            #instTcpSend.REQ := true;
             #instTcpSend.LEN := INT_TO_UDINT(#statSendLenght + 2);

                   IF ((#instTcpSend.DONE)
                       AND (#instTcpSend.BUSY = 0))
                   THEN
                       #instTcpSend.REQ := false;
                       #statStateMQTT := #MQTT_CONNACK;
                       //Delete Send Buffer
                       FOR #statI := 1 TO (#statSendLenght + 2) DO
                           #statSendBuffer[#statI] := 0;
                       END_FOR;
                   ELSIF #instTcpSend.ERROR
                   THEN
                       #statusID := #MQTT_CONNECT;
                       #instTcpSend.REQ := false;
                       #statStateMQTT := #MQTT_ERROR;

                   END_IF;

               END_REGION
               ;
           #MQTT_CONNACK:
               IF #statNewDataRcv THEN

                   IF ((#statRcvBuffer[1] AND b#16#f0) = #MQTT_MSG_TYPE_CONNACK)
                       AND
                       (#statRcvBuffer[4] = #MQTT_CONNACK_ACCEPTED)
                   THEN
                       #statStateMQTT := #MQTT_CONNECTED;
                       #mqttEstablished := true;
                       #busy := false;
                       #statStateMQTTinternal := #IDLE;
                       //start Keep Alive Timer
                       //KeepAliveTImer is set to (Keep Alive (in s) - 2s)
                       #statKeepAliveTime := UINT_TO_TIME((WORD_TO_UINT(#mqttParam.keepAlive) * 1000 - 2000));
                       IF NOT #statKeepAliveOff
                       THEN
                           #statTriggerKeepAlive := true;
                       END_IF;
                       #statNewDataRcv := 0;
                   ELSE
                       #statStateMQTT := #MQTT_ERROR;
                       #statusID := #MQTT_CONNACK;
                   END_IF;
               END_IF;
           #MQTT_CONNECTED:
               IF #publish
                   AND NOT #statPublishOld
                   AND (#statStateMQTTinternal=#IDLE)
               THEN
                   #statStateMQTTinternal := #MQTT_PUBLISH;
                   #published := 0;
                   #error := 0;
                  #statTriggerKeepAlive := false;
                   #statPacketID := #statPacketID + 1;
               END_IF;
               #statPublishOld := #publish;

                IF (#instKeepAlive.Q)
                    AND (#statStateMQTTinternal = #IDLE)
                    AND (NOT #statKeepAliveOff)
                THEN
                    #statStateMQTTinternal := #MQTT_PING;
                    #statTriggerKeepAlive := false;
                END_IF;
                CASE #statStateMQTTinternal OF
                    #IDLE:
                        #published := 0;
                        ;
                    #MQTT_PUBLISH:
                        ;
                        #busy := true;
                        #statConnectLenghtOffset := 0;
                        #statConnectLenght := LEN(IN := #mqttParam.topic) + LEN(IN := #mqttParam.message) + 2;
                        #statSendBuffer[1] := 16#30;
                        #statSendBuffer[1].%X0 := #mqttParam.publishFlag.retain;
                        #statSendBuffer[1].%X3 := false;
                        CASE #mqttParam.publishFlag.qualityOfService OF
                            0:
                                #statSendBuffer[1].%X1 := 0;
                                #statSendBuffer[1].%X2 := 0;
                            1:
                                #statSendBuffer[1].%X1 := 1;
                                #statSendBuffer[1].%X2 := 0;
                                //2 Byte Packet Identifiert added
                                #statConnectLenght := #statConnectLenght + 2;
                            2:
                                #statSendBuffer[1].%X1 := 0;
                                #statSendBuffer[1].%X2 := 1;
                                //2 Byte Packet Identifiert added
                                #statConnectLenght := #statConnectLenght + 2;
                            ELSE:
                                ;
                                #statStateMQTT := #MQTT_ERROR;
                                #statusID := #MQTT_PUBLISH;
                        END_CASE;
                        #statSendLenght := #statConnectLenght;
                        WHILE (#statConnectLenght > 0)
                        DO
                            #statConnectEncodedLenght := #statConnectLenght MOD 128;
                            #statConnectLenght := #statConnectLenght / 128;
                            // if there are more data to encode, set the top bit of this byte
                            IF #statConnectLenght > 0
                            THEN
                                #statConnectEncodedLenght := #statConnectEncodedLenght OR 128;
                                #statSendBuffer[2 + #statConnectLenghtOffset] := INT_TO_BYTE(#statConnectEncodedLenght);
                                #statConnectLenghtOffset := #statConnectLenghtOffset + 1;
                            ELSE
                                #statSendBuffer[2 + #statConnectLenghtOffset] := INT_TO_BYTE(#statConnectEncodedLenght);
                            END_IF;
                        END_WHILE;
                        #statSendLenght := #statSendLenght + #statConnectLenghtOffset;
                        //Variable Header
                        #tempLenght := INT_TO_WORD(LEN(IN := #mqttParam.topic));
                        #statSendBuffer[3 + #statConnectLenghtOffset] := #tempLenght.%B1;
                        #statSendBuffer[4 + #statConnectLenghtOffset] := #tempLenght.%B0;
                        Strg_TO_Chars(Strg := #mqttParam.topic,
                                      pChars := 0,
                                      Cnt => #tempCountChars,
                                      Chars := #tempStringToChar);
                        FOR #statI := 0 TO UINT_TO_INT(#tempCountChars - 1) DO
                            #statSendBuffer[5 + #statConnectLenghtOffset + #statI] := #tempStringToChar[#statI];
                        END_FOR;
                        #statConnectLenghtOffset := #statConnectLenghtOffset + #statI;
                        IF (#mqttParam.publishFlag.qualityOfService > 0)
                        THEN

                            #statSendBuffer[5 + #statConnectLenghtOffset] := #statPacketID.%B1;
                            #statSendBuffer[6 + #statConnectLenghtOffset] := #statPacketID.%B0;
                            //Payload
                            Strg_TO_Chars(Strg := #mqttParam.message,
                                          pChars := 0,
                                          Cnt => #tempCountChars,
                                          Chars := #tempStringToChar);
                            FOR #statI := 0 TO UINT_TO_INT(#tempCountChars - 1) DO
                                #statSendBuffer[7 + #statConnectLenghtOffset + #statI] := #tempStringToChar[#statI];
                            END_FOR;
                            #instTcpSend.LEN := INT_TO_UDINT(#statSendLenght + 2);
                        ELSE
                            Strg_TO_Chars(Strg := #mqttParam.message,
                                          pChars := 0,
                                          Cnt => #tempCountChars,
                                          Chars := #tempStringToChar);
                            FOR #statI := 0 TO UINT_TO_INT(#tempCountChars - 1) DO
                                #statSendBuffer[5 + #statConnectLenghtOffset + #statI] := #tempStringToChar[#statI];
                            END_FOR;
                            #instTcpSend.LEN := INT_TO_UDINT(#statSendLenght + 2);
                        END_IF;

                        #instTcpSend.REQ := true;


                        IF ((#instTcpSend.DONE)
                            AND (#instTcpSend.BUSY = 0))
                        THEN
                            #instTcpSend.REQ := false;
                            IF (#mqttParam.publishFlag.qualityOfService > 0)
                            THEN
                                #statPacketIDAck := #statPacketID;
                                #statStateMQTTinternal := #MQTT_PUBACK;
                            ELSE
                                //QoS = 0; finish here
                                #published := true;
                                #busy := false;
                                #statNewDataRcv := false;
                                IF NOT #statKeepAliveOff
                                THEN
                                    #statTriggerKeepAlive := true;
                                END_IF;

                                #statStateMQTTinternal := #IDLE;
                            END_IF;
                        ELSIF #instTcpSend.ERROR
                        THEN
                            #statusID := #MQTT_PUBLISH;
                            #instTcpSend.REQ := false;
                            #statStateMQTT := #MQTT_ERROR;
                            #status := #instTcpSend.STATUS;
                        END_IF;
                    #MQTT_PUBACK:
                        IF #statNewDataRcv THEN
                            IF ((#statRcvBuffer[1] AND b#16#f0) = #MQTT_MSG_TYPE_PUBACK)
                                OR
                                ((#statRcvBuffer[1] AND b#16#f0) = INT_TO_WORD(#MQTT_MSG_TYPE_PUBREC))
                            THEN
                                IF
                                    (#statRcvBuffer[3] = #statPacketIDAck.%B1)
                                    AND
                                    (#statRcvBuffer[4] = #statPacketIDAck.%B0)
                                THEN
                                    IF (#mqttParam.publishFlag.qualityOfService = 1)
                                    THEN
                                        //QoS = 1; finish here
                                        #statStateMQTTinternal := #MQTT_IDLE;
                                        #published := true;
                                        #busy := false;
                                        #statNewDataRcv := false;
                                        //Re-Activate Kepp Alive Timer
                                        IF NOT #statKeepAliveOff
                                        THEN
                                            #statTriggerKeepAlive := true;
                                        END_IF;

                                        #statStateMQTTinternal := #IDLE;
                                    ELSE
                                        #statStateMQTTinternal := #MQTT_PUBREL;
                                    END_IF;
                                ELSE
                                    #statNewDataRcv := false;
                                END_IF;
                            ELSE
                                #statStateMQTT := #MQTT_ERROR;
                                #statusID := #MQTT_PUBACK;
                            END_IF;
                        END_IF;
                    #MQTT_PUBREL:
                        //fixed Header
                        #statSendBuffer[1] := 16#62;
                        #statSendBuffer[2] := 2;
                        //Variable Header
                        #statSendBuffer[3] := #statPacketID.%B1;
                        #statSendBuffer[4] := #statPacketID.%B0;
                        #instTcpSend.LEN := INT_TO_UDINT(4);
                        #instTcpSend.REQ := true;

                        IF ((#instTcpSend.DONE)
                            AND (#instTcpSend.BUSY = 0))
                        THEN
                            #instTcpSend.REQ := false;
                            #statPacketIDAck := #statPacketID;
                            #statStateMQTTinternal := #MQTT_PUBCOMP;

                        ELSIF #instTcpSend.ERROR
                        THEN
                            #statusID := #MQTT_PUBREL;
                            #instTcpSend.REQ := false;
                            #statStateMQTT := #MQTT_ERROR;
                            #status := #instTcpSend.STATUS;
                        END_IF;
                    #MQTT_PUBCOMP:
                        IF #statNewDataRcv THEN
                            IF ((#statRcvBuffer[1] AND b#16#f0) = #MQTT_MSG_TYPE_PUBCOM)
                            THEN
                                IF
                                    (#statRcvBuffer[3] = #statPacketIDAck.%B1)
                                    AND
                                    (#statRcvBuffer[4] = #statPacketIDAck.%B0)
                                THEN
                                    //QoS = 2; finish here
                                    #statStateMQTTinternal := #MQTT_IDLE;
                                    #published := true;
                                    #busy := false;
                                    #statNewDataRcv := false;
                                    //Re-Activate Kepp Alive Timer
                                    IF NOT #statKeepAliveOff
                                    THEN
                                        #statTriggerKeepAlive := true;
                                    END_IF;

                                    #statStateMQTTinternal := #IDLE;
                                ELSE
                                    #statStateMQTT := #MQTT_ERROR;
                                    #statusID := #MQTT_PUBCOMP;
                                END_IF;
                            END_IF;
                        END_IF;
                    #MQTT_PING:

                        #busy := true;
                        //Build fixed Header
                        //Message Type
                        #statSendBuffer[1] := INT_TO_BYTE(#MQTT_MSG_TYPE_PING);
                        //Remaining Lenght (must be O)
                        #statSendBuffer[2] := 0;
                        #instTcpSend.REQ := true;
                        #instTcpSend.LEN := 2;

                        IF ((#instTcpSend.DONE)
                            AND (#instTcpSend.BUSY = 0))
                        THEN
                            #instTcpSend.REQ := false;
                            #statStateMQTTinternal := #MQTT_PINGRESP;
                        ELSIF #instTcpSend.ERROR
                        THEN
                            #statusID := #MQTT_PING;
                            #instTcpSend.REQ := false;
                            #statStateMQTT := #MQTT_ERROR;
                            #status := #instTcpSend.STATUS;
                        END_IF;
                    #MQTT_PINGRESP:
                        IF #statNewDataRcv
                        THEN
                            IF ((#statRcvBuffer[1] AND b#16#f0) = #MQTT_MSG_TYPE_PINGRESP)
                            THEN
                                #busy := false;
                                #statNewDataRcv := false;
                                #statTriggerKeepAlive := true;
                                #statStateMQTTinternal := #IDLE;
                            END_IF;
                        ELSE
                            #statNewDataRcv := false;
                        END_IF;

                END_CASE;
           #MQTT_DISCONNECT:
           #busy := 0;
           //Build fixed Header
           //Message Type
           #statSendBuffer[1] := INT_TO_BYTE(#MQTT_MSG_TYPE_DISCONNECT);
           //Remaining Lenght (must be O)
           #statSendBuffer[2] := 0;
           #instTcpSend.REQ := true;
           #instTcpSend.LEN := 2;

           IF ((#instTcpSend.DONE)
               AND (#instTcpSend.BUSY = 0))
           THEN
               IF NOT #enable THEN
                   #statStateTCP := #TCP_DISCONNECT;
               END_IF;
               #instTcpSend.REQ := false;
               #statStateMQTT := #MQTT_DISCONNECTED;
               #statStateMQTTinternal := #IDLE;
           ELSIF #instTcpSend.ERROR
           THEN
               IF NOT #enable THEN
                   #statStateTCP := #TCP_DISCONNECT;
               END_IF;
               #statusID := #MQTT_DISCONNECT;
               #instTcpSend.REQ := false;
               #statStateMQTT := #MQTT_ERROR;
               #status := #instTcpSend.STATUS;
           END_IF;
               #MQTT_ERROR:

               REGION Errorhandling MQTT
                   #error := true;
                   #busy := false;
                   #statStateMQTTinternal := #IDLE;
                   #statTriggerKeepAlive := 0;
                   #statKeepAliveOff := false;
                 CASE #statusID OF
                     #MQTT_CONNECT_FLAG_CHECK:
                         #mqttEstablished := false;
                         #statStateMQTT := #MQTT_DISCONNECTED;
                         ;
                     #MQTT_CONNECT:
                         #mqttEstablished := false;
                         #status := #instTcpSend.STATUS;   ;
                         #statStateMQTT := #MQTT_DISCONNECTED;
                       #MQTT_CONNACK:
                           #mqttEstablished := false;
                           #status := #statRcvBuffer[4];
                           #statStateMQTT := #MQTT_DISCONNECTED;
                       #MQTT_PUBLISH:
                               #published := false;
                               #statStateMQTT := #MQTT_CONNECTED;
                               #MQTT_PUBACK,#MQTT_PUBCOMP,#MQTT_PUBREL:
                           #published := false;
                           #status :=#MQTT_ERROR_PACKETID;
                           #statStateMQTT := #MQTT_CONNECTED;
                       #MQTT_PINGRESP:;
                           #MQTT_PING:;
                       #MQTT_DISCONNECT:
                           #mqttEstablished := false;
                          ;
                       ELSE
                           ;
                   END_CASE;
              END_REGION
               ;



       END_CASE
       ;
END_FUNCTION_BLOCK

FUNCTION_BLOCK "FB_MQTT"   // FB5, LAD
{ S7_Optimized_Access := 'TRUE' }
VERSION : 0.1
BEGIN
END_FUNCTION_BLOCK

FUNCTION_BLOCK "FB_concatScrings"   // FB6, LAD
{ S7_Optimized_Access := 'TRUE' }
VERSION : 0.1
   VAR_INPUT
      temperature1 : Real;
      temperature2 : Real;
      temperature3 : Real;
      temperature4 : Real;
      rtd_ch0 : Real;
      rtd_ch1 : Real;
      rtd_ch2 : Real;
      rtd_ch3 : Real;
      presaCounter : UDInt;
      PresaHitrost : Int;
      PresaisRunning : Int;
   END_VAR
   VAR_OUTPUT
      strCombinedString : String;
   END_VAR
   VAR
      tempStr1 : String;
      tempStr2 : String;
      tempStr3 : String;
      tempStr4 : String;
      counterStr : String;
      isRunningStr : String;
      currentSpeedStr : String;
      combinedStr : String;
      rtdStr0 : String;
      rtdStr1 : String;
      rtdStr2 : String;
      rtdStr3 : String;
   END_VAR
BEGIN

REGION Network 2 (SCL)
   // Convert REAL values to STRING
   // 
    VAL_STRG(IN:=#temperature1,
              SIZE:=10,
              PREC:=4,
              FORMAT:=0000,
              P:=16,
              OUT=>#tempStr1);

   //#tempStr1 := REAL_TO_STRING(#temperature1);

     VAL_STRG(IN := #temperature2,
              SIZE := 10,
              PREC := 4,
              FORMAT := 0000,
              P := 16,
              OUT => #tempStr2);

     VAL_STRG(IN := #temperature3,
              SIZE := 10,
              PREC := 4,
              FORMAT := 0000,
              P := 16,
              OUT => #tempStr3);

     VAL_STRG(IN := #temperature4,
              SIZE := 10,
              PREC := 4,
              FORMAT := 0000,
              P := 16,
              OUT => #tempStr4);

   //convert RTD inputs to string
   // Convert RTD values to STRING
   VAL_STRG(IN := #rtd_ch0,
            SIZE := 10,
            PREC := 4,
            FORMAT := 0000,
            P := 16,
            OUT => #rtdStr0);
   VAL_STRG(IN := #rtd_ch1,
            SIZE := 10,
            PREC := 4,
            FORMAT := 0000,
            P := 16,
            OUT => #rtdStr1);
   VAL_STRG(IN := #rtd_ch2,
            SIZE := 10,
            PREC := 4,
            FORMAT := 0000,
            P := 16,
            OUT => #rtdStr2);
   VAL_STRG(IN := #rtd_ch3,
            SIZE := 10,
            PREC := 4,
            FORMAT := 0000,
            P := 16,
            OUT => #rtdStr3);

   // convert int to string
     #currentSpeedStr := ' ';
     VAL_STRG(IN := #PresaHitrost,
              SIZE := 3,
              PREC := 0,
              FORMAT := 0000,
              P := 1,
              OUT => #currentSpeedStr);


   // Convert DINT to STRING
   #counterStr := '';
   VAL_STRG(IN := #presaCounter,
            SIZE := 5,
            PREC := 0,
            FORMAT := 0000,
            P := 1,
            OUT => #counterStr);

   // Convert BOOL to STRING (represent TRUE/FALSE)
   IF #PresaisRunning = 1 THEN
       #isRunningStr := '1';
   ELSE
       #isRunningStr := '0';
   END_IF;

   // Combine all strings into a JSON format
   #combinedStr := '{';
   #combinedStr := CONCAT(IN1 := #combinedStr, IN2 := '"temperature1":');
   #combinedStr := CONCAT(IN1 := #combinedStr, IN2 := #tempStr1);
   #combinedStr := CONCAT(IN1 := #combinedStr, IN2 := ',');
   #combinedStr := CONCAT(IN1 := #combinedStr, IN2 := '"temperature2":');
   #combinedStr := CONCAT(IN1 := #combinedStr, IN2 := #tempStr2);
   #combinedStr := CONCAT(IN1 := #combinedStr, IN2 := ',');
   #combinedStr := CONCAT(IN1 := #combinedStr, IN2 := '"temperature3":');
   #combinedStr := CONCAT(IN1 := #combinedStr, IN2 := #tempStr3);
   #combinedStr := CONCAT(IN1 := #combinedStr, IN2 := ',');
   #combinedStr := CONCAT(IN1 := #combinedStr, IN2 := '"temperature4":');
   #combinedStr := CONCAT(IN1 := #combinedStr, IN2 := #tempStr4);
   #combinedStr := CONCAT(IN1 := #combinedStr, IN2 := ',');

   (* #combinedStr := CONCAT(IN1 := #combinedStr, IN2 := '"rtd_ch0":');
   #combinedStr := CONCAT(IN1 := #combinedStr, IN2 := #rtdStr0);
   #combinedStr := CONCAT(IN1 := #combinedStr, IN2 := ',');

   #combinedStr := CONCAT(IN1 := #combinedStr, IN2 := '"rtd_ch1":');
   #combinedStr := CONCAT(IN1 := #combinedStr, IN2 := #rtdStr1);
   #combinedStr := CONCAT(IN1 := #combinedStr, IN2 := ',');
   *)
   #combinedStr := CONCAT(IN1 := #combinedStr, IN2 := '"rtd_ch2":');
   #combinedStr := CONCAT(IN1 := #combinedStr, IN2 := #rtdStr2);
   #combinedStr := CONCAT(IN1 := #combinedStr, IN2 := ',');


   #combinedStr := CONCAT(IN1 := #combinedStr, IN2 := '"counter":');
   #combinedStr := CONCAT(IN1 := #combinedStr, IN2 := #counterStr);
   #combinedStr := CONCAT(IN1 := #combinedStr, IN2 := ',');
   #combinedStr := CONCAT(IN1 := #combinedStr, IN2 := '"isRunning":');
   #combinedStr := CONCAT(IN1 := #combinedStr, IN2 := #isRunningStr);
   #combinedStr := CONCAT(IN1 := #combinedStr, IN2 := ',');
   #combinedStr := CONCAT(IN1 := #combinedStr, IN2 := '"currentSpeed":');
   #combinedStr := CONCAT(IN1 := #combinedStr, IN2 := #currentSpeedStr);
   #combinedStr := CONCAT(IN1 := #combinedStr, IN2 := '}');

   // Now combinedStr contains the concatenated string in JSON format
   #strCombinedString := #combinedStr;
END_REGION
END_FUNCTION_BLOCK

FUNCTION_BLOCK "FB_CONCAT_STRINGS_FOR_MQTT"   // FB7, LAD
{ S7_Optimized_Access := 'TRUE' }
VERSION : 0.1
   VAR_INPUT
      temperature1 : Real;
      temperature2 : Real;
      temperature3 : Real;
      temperature4 : Real;
   END_VAR
   VAR_OUTPUT
      strCombinedString : String;
      q_aStringToSendToMqtt : Array[0..1] of String;
   END_VAR
   VAR
      tempStr1 : String;
      tempStr2 : String;
      tempStr3 : String;
      tempStr4 : String;
      combinedStr : String;
      lenghtOfCombinedString : Int;
      Static_1 : Int;
      assocValues : Array[0..3] of DInt;
      combineStr_1 : String;
      combineStr_2 : String;
   END_VAR
BEGIN

REGION Network 2 (SCL)
   // Convert REAL values to STRING
   // 
   VAL_STRG(IN := #temperature1,
            SIZE := 10,
            PREC := 4,
            FORMAT := 0000,
            P := 16,
            OUT => #tempStr1);

   //#tempStr1 := REAL_TO_STRING(#temperature1);

   VAL_STRG(IN := #temperature2,
            SIZE := 10,
            PREC := 4,
            FORMAT := 0000,
            P := 16,
            OUT => #tempStr2);

   VAL_STRG(IN := #temperature3,
            SIZE := 10,
            PREC := 4,
            FORMAT := 0000,
            P := 16,
            OUT => #tempStr3);

   VAL_STRG(IN := #temperature4,
            SIZE := 10,
            PREC := 4,
            FORMAT := 0000,
            P := 16,
            OUT => #tempStr4);


   // Combine all strings into a JSON format
   #combinedStr := '{';
   #combinedStr := CONCAT(IN1 := #combinedStr, IN2 := '"temperature1":');
   #combinedStr := CONCAT(IN1 := #combinedStr, IN2 := #tempStr1);
   #combinedStr := CONCAT(IN1 := #combinedStr, IN2 := ',');
   #combinedStr := CONCAT(IN1 := #combinedStr, IN2 := '"temperature2":');
   #combinedStr := CONCAT(IN1 := #combinedStr, IN2 := #tempStr2);
   #combinedStr := CONCAT(IN1 := #combinedStr, IN2 := ',');
   #combinedStr := CONCAT(IN1 := #combinedStr, IN2 := '"temperature3":');
   #combinedStr := CONCAT(IN1 := #combinedStr, IN2 := #tempStr3);
   #combinedStr := CONCAT(IN1 := #combinedStr, IN2 := ',');
   #combinedStr := CONCAT(IN1 := #combinedStr, IN2 := '"temperature4":');
   #combinedStr := CONCAT(IN1 := #combinedStr, IN2 := #tempStr4);
   #combinedStr := CONCAT(IN1 := #combinedStr, IN2 := '}');

   // Now combinedStr contains the concatenated string in JSON format
   #strCombinedString := #combinedStr;

   #lenghtOfCombinedString := LEN(#combinedStr);


   // Check if the length exceeds 254 characters
   IF #lenghtOfCombinedString > 254 THEN
       // Extract the first 254 characters for combineStr_1
       #combineStr_1 := LEFT(IN := #combinedStr, L := 254);

       // Extract the remaining characters for combineStr_2
       #combineStr_2 := RIGHT(IN := #combinedStr, L := #lenghtOfCombinedString - 254);
   ELSE
       // If length is less than or equal to 254, use the entire string in combineStr_1
       #combineStr_1 := #combinedStr;
       #combineStr_2 := '';  // Set combineStr_2 to an empty string
   END_IF;

   #q_aStringToSendToMqtt[0] := #combineStr_1;
   #q_aStringToSendToMqtt[1] := #combineStr_2;
END_REGION
END_FUNCTION_BLOCK

FUNCTION_BLOCK "FB_CONCAT_STRINGS_FOR_MQTT_1"   // FB9, LAD
{ S7_Optimized_Access := 'TRUE' }
VERSION : 0.1
   VAR_INPUT
      temperature1 : Real;
      temperature2 : Real;
      temperature3 : Real;
      temperature4 : Real;
      customText : String;
   END_VAR
   VAR_OUTPUT
      strCombinedString : String;
      q_aStringToSendToMqtt : Array[0..1] of String;
   END_VAR
   VAR
      tempStr1 : String;
      tempStr2 : String;
      tempStr3 : String;
      tempStr4 : String;
      combinedStr : String;
      lenghtOfCombinedString : Int;
      Static_1 : Int;
      assocValues : Array[0..3] of DInt;
      combineStr_1 : String;
      combineStr_2 : String;
      currentStrLength : Int;
      tempStrLength : Int;
      SafeConcat : "FB_saveConcat";
   END_VAR
BEGIN

REGION Network 2 (SCL)
   // Initialize variables
   #combinedStr := '{';
   #combineStr_1 := ''; // First part of the JSON
   #combineStr_2 := ''; // Second part of the JSON

   // Convert REAL values to STRING
   VAL_STRG(IN := #temperature1,
            SIZE := 10,
            PREC := 4,
            FORMAT := 0000,
            P := 16,
            OUT => #tempStr1);

   VAL_STRG(IN := #temperature2,
            SIZE := 10,
            PREC := 4,
            FORMAT := 0000,
            P := 16,
            OUT => #tempStr2);

   VAL_STRG(IN := #temperature3,
            SIZE := 10,
            PREC := 4,
            FORMAT := 0000,
            P := 16,
            OUT => #tempStr3);

   VAL_STRG(IN := #temperature4,
            SIZE := 10,
            PREC := 4,
            FORMAT := 0000,
            P := 16,
            OUT => #tempStr4);

   // Start constructing the JSON string

   // Concatenate temperature1
   #SafeConcat(IN1 := #customText,
               IN2 := #tempStr1,
               combineStr_1 := #combineStr_1,
               combineStr_2 := #combineStr_2,
               SafeConcat => #combinedStr);

   #SafeConcat(IN1 := ',',
               IN2 := '',
               combineStr_1 := #combineStr_1,
               combineStr_2 := #combineStr_2,
               SafeConcat => #combinedStr);

   // Concatenate temperature2
   #SafeConcat(IN1 := '"temperature2":',
               IN2 := #tempStr2,
               combineStr_1 := #combineStr_1,
               combineStr_2 := #combineStr_2,
               SafeConcat => #combinedStr);

   #SafeConcat(IN1 := ',',
               IN2 := '',
               combineStr_1 := #combineStr_1,
               combineStr_2 := #combineStr_2,
               SafeConcat => #combinedStr);

   // Concatenate temperature3
   #SafeConcat(IN1 := '"temperature3":',
               IN2 := #tempStr3,
               combineStr_1 := #combineStr_1,
               combineStr_2 := #combineStr_2,
               SafeConcat => #combinedStr);

   #SafeConcat(IN1 := ',',
               IN2 := '',
               combineStr_1 := #combineStr_1,
               combineStr_2 := #combineStr_2,
               SafeConcat => #combinedStr);

   // Concatenate temperature4
   #SafeConcat(IN1 := '"temperature4":',
               IN2 := #tempStr4,
               combineStr_1 := #combineStr_1,
               combineStr_2 := #combineStr_2,
               SafeConcat => #combinedStr);

   #SafeConcat(IN1 := '}',
               IN2 := '',
               combineStr_1 := #combineStr_1,
               combineStr_2 := #combineStr_2,
               SafeConcat => #combinedStr);

   // Now #combineStr_1 and #combineStr_2 hold the JSON formatted string, split if necessary
   #q_aStringToSendToMqtt[0] := #combineStr_1;
   #q_aStringToSendToMqtt[1] := #combineStr_2;
   #lenghtOfCombinedString := LEN(IN:=#q_aStringToSendToMqtt[0]) + LEN(IN:=#q_aStringToSendToMqtt[1]);
END_REGION
END_FUNCTION_BLOCK

FUNCTION_BLOCK "FB_saveConcat"   // FB10, LAD
{ S7_Optimized_Access := 'TRUE' }
VERSION : 0.1
   VAR_INPUT
      IN1 : String;
      IN2 : String;
   END_VAR
   VAR_OUTPUT
      SafeConcat : String;
   END_VAR
   VAR_IN_OUT
      combineStr_1 : String;
      combineStr_2 : String;
   END_VAR
   VAR
      tempStrLength : Int;
   END_VAR
BEGIN

REGION Network 2 (SCL)

   #tempStrLength :=LEN(#combineStr_1) + LEN(#IN1) + LEN(#IN2);
   IF #tempStrLength <= 254 THEN
       // Safe to concatenate and store in #combineStr_1
       #SafeConcat := CONCAT(IN1 := #IN1, IN2 := #IN2);
       #combineStr_1 := CONCAT(IN1:=#combineStr_1, IN2 := #SafeConcat);
   ELSE
       #SafeConcat := CONCAT(IN1 := #IN1, IN2 := #IN2);
       #combineStr_2 := CONCAT(IN1 := #combineStr_2, IN2 := #SafeConcat);

   END_IF;
END_REGION
END_FUNCTION_BLOCK

FUNCTION_BLOCK "FB_ServoGo"   // FB12, LAD
{ S7_Optimized_Access := 'TRUE' }
VERSION : 0.1
BEGIN
END_FUNCTION_BLOCK

FUNCTION_BLOCK "PTC_1000_resistanceCalculation"   // FB13, LAD
{ S7_Optimized_Access := 'TRUE' }
VERSION : 0.1
   VAR_INPUT
      Coeff1 : Real;
      Coeff2 : Real;
      coeff3 : Real;
      constat : Real;
      PTC_resistance : DInt;
   END_VAR
   VAR_OUTPUT
      q_rTemp : Real;
   END_VAR
   VAR
      _rt_r25 : Real;
      _temperature : Real;
   END_VAR
BEGIN

REGION Network 2 (SCL)

   #_rt_r25 := #PTC_resistance / 1000.0;
   #_temperature := (#coeff3 * #_rt_r25 ** 3) + (#Coeff2 * #_rt_r25 ** 2) + (#Coeff1 * #_rt_r25) + #constat;

   #q_rTemp := #_temperature;
END_REGION
END_FUNCTION_BLOCK

FUNCTION_BLOCK "FB_EgasiMotorControl"   // FB16, LAD
{ S7_Optimized_Access := 'TRUE' }
VERSION : 0.1
   VAR_INPUT
      i_xPWR_48 : Bool;
      i_xInPOS1 : Bool;
      i_xInPOS2 : Bool;
      i_xisHommed : Bool;
      i_xExternalError : Bool;
      i_xDemoPeriod : Bool;
      i_wRawTempValue : Word;
      i_xGoPOS1_Automatic : Bool;
      i_xGOPOS2_Automatic : Bool;
      i_rCurrentRawMINValue : Real;
      i_rCurrentRawMAXValue : Real;
      i_HMIxOverRideControl : Bool;
      i_xHMI_demoMode : Bool;   // Clock 1Hz
      i_xHMI_automaticMode : Bool;   // Automatic Mode for production
   END_VAR
   VAR_OUTPUT
      q_xMotorPWR : Bool;
      q_xGoPOS1 : Bool;
      q_xGoPOS2 : Bool;
      q_xGoHOME : Bool;
      q_rScaledTemperature : Real;
      q_xErrorPOS1 : Bool;
      q_xErrorPOS2 : Bool;
      q_xFuseERR : Bool;
      q_xMotorERR : Bool;
      q_xinPOS1 : Bool;
      q_xInPOS2 : Bool;
   END_VAR
   VAR_IN_OUT
      io_HMI_data : "UDT_MotorControl";
      UDT_EGASI : "EGASI_MOTOR_CONTROL";
   END_VAR
   VAR
      POS1_timer : TON_TIME;
      POS2_timer : TON_TIME;
      DemoClock : Bool;
      HW_RESET_PULSE : TP_TIME;
   END_VAR
   VAR RETAIN
      pulsemerker : Bool;
      s_HMI_gopos1 : Bool;
   END_VAR
   VAR
      s_HMI_gopos2 : Bool;
   END_VAR
   VAR RETAIN
      s_bits : Array[0..3] of Bool;
      xIncrementbits : Bool;
      Counter_POS1 : UDInt;
      Counter_POS2 : UDInt;
   END_VAR
   VAR_TEMP
      bits : Array[0..2] of Bool;
   END_VAR
   VAR_TEMP   // added for the SCL form of the ladder/FBD networks
      _w1 : Bool;
      _w2 : Bool;
      _w3 : Bool;
      _w4 : Bool;
   END_VAR
BEGIN

REGION Network 1: EGASI UDT CONTROL -> MAPPING UDT DB
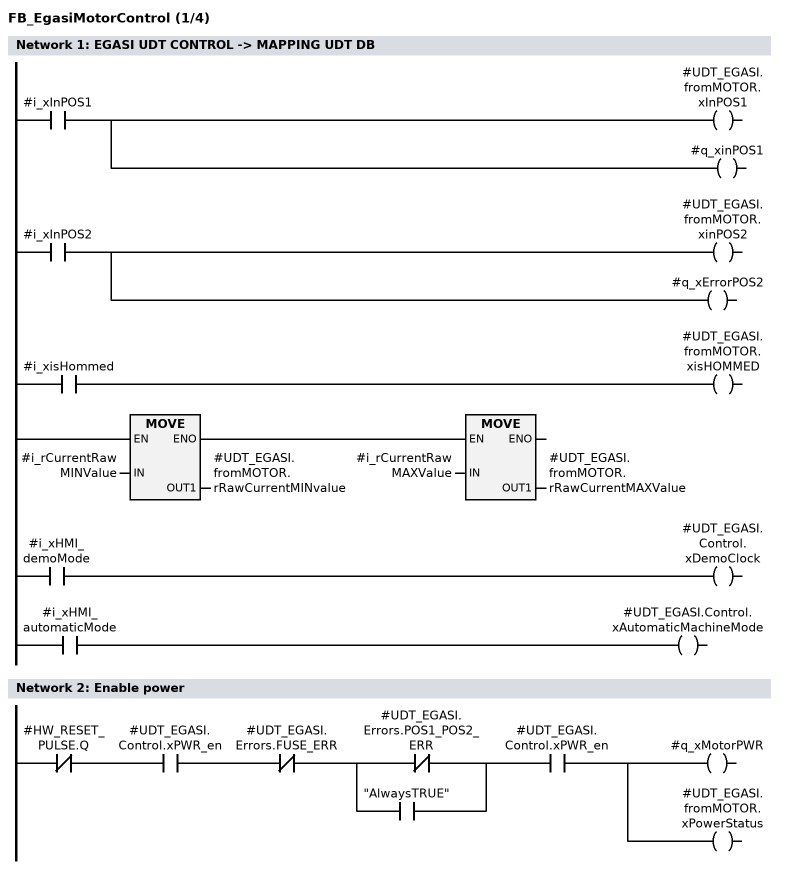
   RUNG wire#powerrail
      Contact( #i_xInPOS1 )
      wire#w1
      Coil( #UDT_EGASI.fromMOTOR.xInPOS1 )
   END_RUNG
   RUNG wire#w1
      Coil( #q_xinPOS1 )
   END_RUNG
   RUNG wire#powerrail
      Contact( #i_xInPOS2 )
      wire#w2
      Coil( #UDT_EGASI.fromMOTOR.xinPOS2 )
   END_RUNG
   RUNG wire#w2
      Coil( #q_xErrorPOS2 )
   END_RUNG
   RUNG wire#powerrail
      Contact( #i_xisHommed )
      Coil( #UDT_EGASI.fromMOTOR.xisHOMMED )
   END_RUNG
   RUNG wire#powerrail
      Move(in := #i_rCurrentRawMINValue, out1 => #UDT_EGASI.fromMOTOR.rRawCurrentMINvalue)
      Move(in := #i_rCurrentRawMAXValue, out1 => #UDT_EGASI.fromMOTOR.rRawCurrentMAXValue)
   END_RUNG
   RUNG wire#powerrail
      Contact( #i_xHMI_demoMode )
      Coil( #UDT_EGASI.Control.xDemoClock )
   END_RUNG
   RUNG wire#powerrail
      Contact( #i_xHMI_automaticMode )
      Coil( #UDT_EGASI.Control.xAutomaticMachineMode )
   END_RUNG
   // the same network as SCL:
   #UDT_EGASI.fromMOTOR.xInPOS1 := #i_xInPOS1;
   #q_xinPOS1 := #i_xInPOS1;
   #UDT_EGASI.fromMOTOR.xinPOS2 := #i_xInPOS2;
   #q_xErrorPOS2 := #i_xInPOS2;
   #UDT_EGASI.fromMOTOR.xisHOMMED := #i_xisHommed;
   #UDT_EGASI.fromMOTOR.rRawCurrentMINvalue := #i_rCurrentRawMINValue;
   #UDT_EGASI.fromMOTOR.rRawCurrentMAXValue := #i_rCurrentRawMAXValue;
   #UDT_EGASI.Control.xDemoClock := #i_xHMI_demoMode;
   #UDT_EGASI.Control.xAutomaticMachineMode := #i_xHMI_automaticMode;
END_REGION

REGION Network 2: Enable power
   RUNG wire#powerrail
      I_Contact( #HW_RESET_PULSE.Q )
      Contact( #UDT_EGASI.Control.xPWR_en )
      I_Contact( #UDT_EGASI.Errors.FUSE_ERR )
      wire#w1
      I_Contact( #UDT_EGASI.Errors.POS1_POS2_ERR )
      wire#w2
      Contact( #UDT_EGASI.Control.xPWR_en )
      wire#w3
      Coil( #q_xMotorPWR )
   END_RUNG
   RUNG wire#w1
      Contact( "AlwaysTRUE" )
   END_RUNG wire#w2
   RUNG wire#w3
      Coil( #UDT_EGASI.fromMOTOR.xPowerStatus )
   END_RUNG
   // the same network as SCL:
   #q_xMotorPWR := NOT #HW_RESET_PULSE.Q AND #UDT_EGASI.Control.xPWR_en AND NOT #UDT_EGASI.Errors.FUSE_ERR AND (NOT #UDT_EGASI.Errors.POS1_POS2_ERR OR "AlwaysTRUE") AND #UDT_EGASI.Control.xPWR_en;
   #UDT_EGASI.fromMOTOR.xPowerStatus := #q_xMotorPWR;
END_REGION

REGION Network 3: Position control
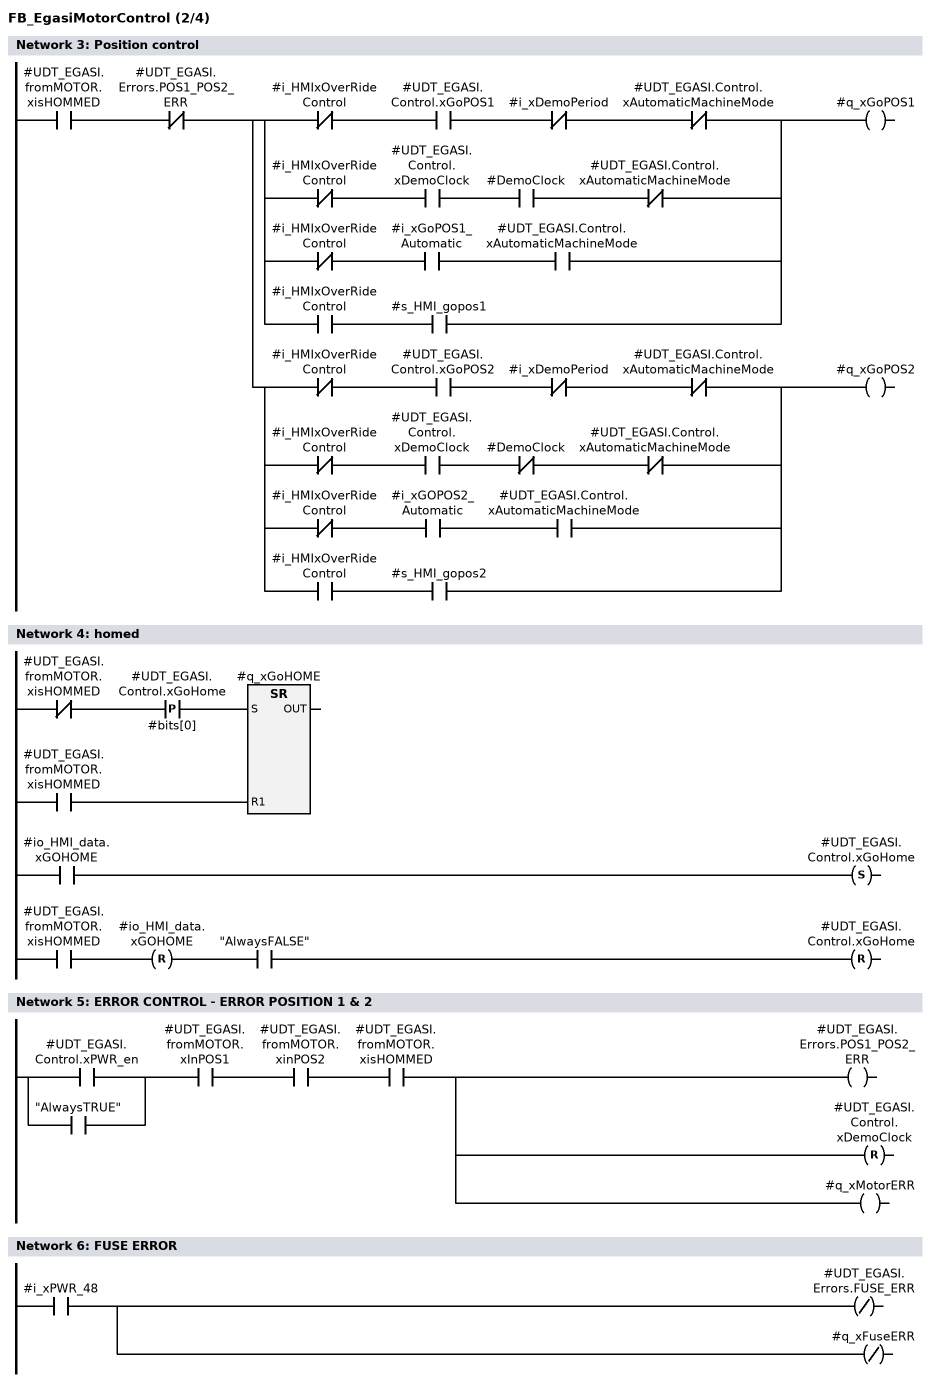
   RUNG wire#powerrail
      Contact( #UDT_EGASI.fromMOTOR.xisHOMMED )
      I_Contact( #UDT_EGASI.Errors.POS1_POS2_ERR )
      wire#w1
      I_Contact( #i_HMIxOverRideControl )
      Contact( #UDT_EGASI.Control.xGoPOS1 )
      I_Contact( #i_xDemoPeriod )
      I_Contact( #UDT_EGASI.Control.xAutomaticMachineMode )
      wire#w2
      Coil( #q_xGoPOS1 )
   END_RUNG
   RUNG wire#w1
      I_Contact( #i_HMIxOverRideControl )
      Contact( #UDT_EGASI.Control.xDemoClock )
      Contact( #DemoClock )
      I_Contact( #UDT_EGASI.Control.xAutomaticMachineMode )
   END_RUNG wire#w2
   RUNG wire#w1
      I_Contact( #i_HMIxOverRideControl )
      Contact( #i_xGoPOS1_Automatic )
      Contact( #UDT_EGASI.Control.xAutomaticMachineMode )
   END_RUNG wire#w2
   RUNG wire#w1
      Contact( #i_HMIxOverRideControl )
      Contact( #s_HMI_gopos1 )
   END_RUNG wire#w2
   RUNG wire#w1
      I_Contact( #i_HMIxOverRideControl )
      Contact( #UDT_EGASI.Control.xGoPOS2 )
      I_Contact( #i_xDemoPeriod )
      I_Contact( #UDT_EGASI.Control.xAutomaticMachineMode )
      wire#w3
      Coil( #q_xGoPOS2 )
   END_RUNG
   RUNG wire#w1
      I_Contact( #i_HMIxOverRideControl )
      Contact( #UDT_EGASI.Control.xDemoClock )
      I_Contact( #DemoClock )
      I_Contact( #UDT_EGASI.Control.xAutomaticMachineMode )
   END_RUNG wire#w3
   RUNG wire#w1
      I_Contact( #i_HMIxOverRideControl )
      Contact( #i_xGOPOS2_Automatic )
      Contact( #UDT_EGASI.Control.xAutomaticMachineMode )
   END_RUNG wire#w3
   RUNG wire#w1
      Contact( #i_HMIxOverRideControl )
      Contact( #s_HMI_gopos2 )
   END_RUNG wire#w3
   // the same network as SCL:
   #_w1 := #UDT_EGASI.fromMOTOR.xisHOMMED AND NOT #UDT_EGASI.Errors.POS1_POS2_ERR;
   #q_xGoPOS1 := #_w1 AND ((NOT #i_HMIxOverRideControl AND #UDT_EGASI.Control.xGoPOS1 AND NOT #i_xDemoPeriod AND NOT #UDT_EGASI.Control.xAutomaticMachineMode) OR (NOT #i_HMIxOverRideControl AND #UDT_EGASI.Control.xDemoClock AND #DemoClock AND NOT #UDT_EGASI.Control.xAutomaticMachineMode) OR (NOT #i_HMIxOverRideControl AND #i_xGoPOS1_Automatic AND #UDT_EGASI.Control.xAutomaticMachineMode) OR (#i_HMIxOverRideControl AND #s_HMI_gopos1));
   #q_xGoPOS2 := #_w1 AND ((NOT #i_HMIxOverRideControl AND #UDT_EGASI.Control.xGoPOS2 AND NOT #i_xDemoPeriod AND NOT #UDT_EGASI.Control.xAutomaticMachineMode) OR (NOT #i_HMIxOverRideControl AND #UDT_EGASI.Control.xDemoClock AND NOT #DemoClock AND NOT #UDT_EGASI.Control.xAutomaticMachineMode) OR (NOT #i_HMIxOverRideControl AND #i_xGOPOS2_Automatic AND #UDT_EGASI.Control.xAutomaticMachineMode) OR (#i_HMIxOverRideControl AND #s_HMI_gopos2));
END_REGION

REGION Network 4: homed
   RUNG wire#powerrail
      I_Contact( #UDT_EGASI.fromMOTOR.xisHOMMED )
      P_Contact(operand := #UDT_EGASI.Control.xGoHome, bit := #bits[0])
      S_SR(operand := #q_xGoHOME, r1 := wire#w1)
   END_RUNG
   RUNG wire#powerrail
      Contact( #UDT_EGASI.fromMOTOR.xisHOMMED )
   END_RUNG wire#w1
   RUNG wire#powerrail
      Contact( #io_HMI_data.xGOHOME )
      S_Coil( #UDT_EGASI.Control.xGoHome )
   END_RUNG
   RUNG wire#powerrail
      Contact( #UDT_EGASI.fromMOTOR.xisHOMMED )
      R_Coil( #io_HMI_data.xGOHOME )
      Contact( "AlwaysFALSE" )
      R_Coil( #UDT_EGASI.Control.xGoHome )
   END_RUNG
   // the same network as SCL:
   #_w1 := NOT #UDT_EGASI.fromMOTOR.xisHOMMED AND #UDT_EGASI.Control.xGoHome AND NOT #bits[0];   // rising edge of #UDT_EGASI.Control.xGoHome
   #bits[0] := #UDT_EGASI.Control.xGoHome;
   IF #_w1 THEN
       #q_xGoHOME := TRUE;   // SR flip-flop
   END_IF;
   IF #UDT_EGASI.fromMOTOR.xisHOMMED THEN #q_xGoHOME := FALSE; END_IF;
   IF #io_HMI_data.xGOHOME THEN #UDT_EGASI.Control.xGoHome := TRUE; END_IF;
   IF #UDT_EGASI.fromMOTOR.xisHOMMED THEN #io_HMI_data.xGOHOME := FALSE; END_IF;
   IF #UDT_EGASI.fromMOTOR.xisHOMMED AND "AlwaysFALSE" THEN #UDT_EGASI.Control.xGoHome := FALSE; END_IF;
END_REGION

REGION Network 5: ERROR CONTROL - ERROR POSITION 1 & 2
   RUNG wire#powerrail
      Contact( #UDT_EGASI.Control.xPWR_en )
      wire#w1
      Contact( #UDT_EGASI.fromMOTOR.xInPOS1 )
      Contact( #UDT_EGASI.fromMOTOR.xinPOS2 )
      Contact( #UDT_EGASI.fromMOTOR.xisHOMMED )
      wire#w2
      Coil( #UDT_EGASI.Errors.POS1_POS2_ERR )
   END_RUNG
   RUNG wire#powerrail
      Contact( "AlwaysTRUE" )
   END_RUNG wire#w1
   RUNG wire#w2
      R_Coil( #UDT_EGASI.Control.xDemoClock )
   END_RUNG
   RUNG wire#w2
      Coil( #q_xMotorERR )
   END_RUNG
   // the same network as SCL:
   #UDT_EGASI.Errors.POS1_POS2_ERR := (#UDT_EGASI.Control.xPWR_en OR "AlwaysTRUE") AND #UDT_EGASI.fromMOTOR.xInPOS1 AND #UDT_EGASI.fromMOTOR.xinPOS2 AND #UDT_EGASI.fromMOTOR.xisHOMMED;
   IF #UDT_EGASI.Errors.POS1_POS2_ERR THEN #UDT_EGASI.Control.xDemoClock := FALSE; END_IF;
   #q_xMotorERR := #UDT_EGASI.Errors.POS1_POS2_ERR;
END_REGION

REGION Network 6: FUSE ERROR
   RUNG wire#powerrail
      Contact( #i_xPWR_48 )
      wire#w1
      I_Coil( #UDT_EGASI.Errors.FUSE_ERR )
   END_RUNG
   RUNG wire#w1
      I_Coil( #q_xFuseERR )
   END_RUNG
   // the same network as SCL:
   #UDT_EGASI.Errors.FUSE_ERR := NOT #i_xPWR_48;
   #q_xFuseERR := NOT #i_xPWR_48;
END_REGION

REGION Network 7: POSITION ERROR POS1